VERSION : 0.1
   VAR
      General : Struct
         ManipulatorFaultProximitiSwitch : Bool;
         ManipulatorFaultRuntime : Bool;
         CPCleanerFaultProximitiSwitch : Bool;
         CPCleanerFaultRuntime : Bool;
         PCPCleaner : Bool;
         Spare6 : Bool;
         Spare7 : Bool;
         Spare8 : Bool;
         Spare9 : Bool;
         Spare10 : Bool;
         Spare11 : Bool;
         Spare12 : Bool;
         Spare13 : Bool;
         Spare14 : Bool;
         Spare15 : Bool;
         Spare16 : Bool;
      END_STRUCT;
      SafteyDeviceSelected : Array[1..16] of Bool;
      "Saftey DeviceAS" : Array[1..16] of Bool;   // Automatic stop at the Saftey Device
      "Saftey DeviceES" : Array[1..16] of Bool;   // Emergency stop at the Saftey Device
   END_VAR
BEGIN
END_DATA_BLOCK

DATA_BLOCK "DB1031_AddStatus"   // DB1031
{ S7_Optimized_Access := 'FALSE' }
VERSION : 0.1
   VAR
      SaftyDevice : Array[0..4] of "UDT_SafetyDevice";
   END_VAR
BEGIN
END_DATA_BLOCK

DATA_BLOCK "DB1040_TT_MovementFault"   // DB1040
{ S7_Optimized_Access := 'FALSE' }
VERSION : 0.1
   VAR
      General : Struct
         MLD_Taktdehnung1Aktiv : Bool;   // Taktdehnung 01 ist aktiv
         MLD_Taktdehnung2Aktiv : Bool;   // Taktdehnung 02 ist aktiv
         MLD_Taktdehnung3Aktiv : Bool;   // Taktdehnung 03 ist aktiv
         MLD_Taktdehnung4Aktiv : Bool;   // Taktdehnung 04 ist aktiv
         STG_Reserve_0_4 : Bool;
         STG_Reserve_0_5 : Bool;
         STG_Reserve_0_6 : Bool;
         STG_Reserve_0_7 : Bool;
         STG_Reserve_1_0 : Bool;
         STG_Reserve_1_1 : Bool;
         STG_Reserve_1_2 : Bool;
         STG_Reserve_1_3 : Bool;
         STG_Reserve_1_4 : Bool;
         STG_Reserve_1_5 : Bool;
         STG_Reserve_1_6 : Bool;
         STG_Reserve_1_7 : Bool;
      END_STRUCT;
      IPOS : Struct
         STG_Luefter : Bool;   // Störung Grp2: Der Versorgung oder des Motorschutzes des Lüfters
         STG_Umrichter : Bool;   // Störung: Der Umrichter ist nicht betriebsbereit
         STG_Motorschutz : Bool;   // Störung: Der Versorgung oder des Motorschutzes des Umrichters
         STG_von_IPOS : Bool;   // Störung: Ein Störungssignal von dem Umrichter steht an
         STG_Genauhaltini : Bool;   // Störung: Die Genauhalteposition (Initiator) wurde nicht erreicht
         STG_Genauhalt_immer_ein : Bool;   // Störung: Die Genauhalteposition (Initiator) wird dauernd belegt
         STG_Busfehler : Bool;   // Störung: Busteilnehmer ist nicht erreichbar
         STG_Reserve_0_7 : Bool;
         STG_Reserve_1_0 : Bool;
         STG_Reserve_1_1 : Bool;
         STG_Reserve_1_2 : Bool;
         STG_Reserve_1_3 : Bool;
         STG_Reserve_1_4 : Bool;
         STG_Reserve_1_5 : Bool;
         STG_Reserve_1_6 : Bool;
         STG_Reserve_1_7 : Bool;
      END_STRUCT;
      Segmentkennung : Struct
         STG_Nummer_unlogisch : Bool;
         STG_Hardwareabschaltung : Bool;
         STG_Wechsel_in_Pos : Bool;
         STG_Reserve_0_3 : Bool;
         STG_Reserve_0_4 : Bool;
         STG_Reserve_0_5 : Bool;
         STG_Reserve_0_6 : Bool;
         STG_Reserve_0_7 : Bool;
         STG_Reserve_1_0 : Bool;
         STG_Reserve_1_1 : Bool;
         STG_Reserve_1_2 : Bool;
         STG_Reserve_1_3 : Bool;
         STG_Reserve_1_4 : Bool;
         STG_Reserve_1_5 : Bool;
         STG_Reserve_1_6 : Bool;
         STG_Reserve_1_7 : Bool;
      END_STRUCT;
      Kettenspanner : Struct
         STG_Entlastung : Bool;
         STG_Druckaufbau : Bool;
         STG_Reserve_0_2 : Bool;
         STG_Reserve_0_3 : Bool;
         STG_Reserve_0_4 : Bool;
         STG_Reserve_0_5 : Bool;
         STG_Reserve_0_6 : Bool;
         STG_Reserve_0_7 : Bool;
         STG_Reserve_1_0 : Bool;
         STG_Reserve_1_1 : Bool;
         STG_Reserve_1_2 : Bool;
         STG_Reserve_1_3 : Bool;
         STG_Reserve_1_4 : Bool;
         STG_Reserve_1_5 : Bool;
         STG_Reserve_1_6 : Bool;
         STG_Reserve_1_7 : Bool;
      END_STRUCT;
   END_VAR
BEGIN
END_DATA_BLOCK

DATA_BLOCK "DB1049_TT_Value"   // DB1049
{ S7_Optimized_Access := 'FALSE' }
AUTHOR : KT242
VERSION : 0.1
   VAR
      Taktzeit : S5Time := S5T#15S;
      Vorwarnzeit : S5Time := S5T#1S;
      Seg_fuer_WW : Int := 0;
      Seg_fuer_Teachen : Int := 0;
      Pos_Offset_Stop : Int := 0;
      Pos_Offset_WW : Int := 0;
      Pos_Offset_Teachen : Int := 0;
      Antrieb_RP : Int := 5000;
      Antrieb_RN : Int := 5000;
      Antrieb_Hand : Int := 500;
      Antrieb_Auto : Int := 1200;
      WaitTimeMHFront : S5Time := S5T#2S;
      RunTimeManipulator : S5Time := S5T#30S;
      RunTimeCPCleaner : S5Time := S5T#5S;
      DelayTimeCPCleaning : S5Time := S5T#500MS;
      DurationCPCleaning : S5Time := S5T#2S;
   END_VAR
BEGIN
END_DATA_BLOCK

DATA_BLOCK "DB1050_Seg_Fault"   // DB1050
{ S7_Optimized_Access := 'FALSE' }
VERSION : 0.1
   VAR
      General : Struct
         STG_Reserve_0_0 : Bool;
         STG_Reserve_0_1 : Bool;
         STG_Reserve_0_2 : Bool;
         STG_Reserve_0_3 : Bool;
         STG_Reserve_0_4 : Bool;
         STG_Reserve_0_5 : Bool;
         STG_Reserve_0_6 : Bool;
         STG_Reserve_0_7 : Bool;
         STG_Reserve_1_0 : Bool;
         STG_Reserve_1_1 : Bool;
         STG_Reserve_1_2 : Bool;
         STG_Reserve_1_3 : Bool;
         STG_Reserve_1_4 : Bool;
         STG_Reserve_1_5 : Bool;
         STG_Reserve_1_6 : Bool;
         STG_Reserve_1_7 : Bool;
      END_STRUCT;
      Segmentverwaltung : Struct
         STG_keine_SegmentNr : Bool;   // Störung Grp3: Es ist keine Segmentkennung vorhanden
         STG_falsche_Paritaet : Bool;   // Störung Grp1: Das Paritätsbit wurde falsch gesetzt
         STG_SegNr_zu_gross : Bool;   // Störung Grp1: Die verdrahtete Segmentnummer ist für dieses RT zu Groß
         STG_Platz_doppelt : Bool;   // Störung Grp1: der Platz auf dem Segment wurde doppelt belegt // Verdrahtungsfehler
         STG_Reserve_0_4 : Bool;
         STG_Reserve_0_5 : Bool;
         STG_Reserve_0_6 : Bool;
         STG_Reserve_0_7 : Bool;
         STG_Reserve_1_0 : Bool;
         STG_Reserve_1_1 : Bool;
         STG_Reserve_1_2 : Bool;
         STG_Reserve_1_3 : Bool;
         STG_Reserve_1_4 : Bool;
         STG_Reserve_1_5 : Bool;
         STG_Reserve_1_6 : Bool;
         STG_Reserve_1_7 : Bool;
      END_STRUCT;
   END_VAR
BEGIN
END_DATA_BLOCK

DATA_BLOCK "DB1051_TT_SegValue"   // DB1051
{ S7_Optimized_Access := 'FALSE' }
VERSION : 0.1
   VAR
      Station : Array[1..8] of Struct
         FoamingEnable : Bool;
         MovingEnable : Bool;
         ToolChange : Bool;
         Spare4 : Bool;
         Spare5 : Bool;
         Spare6 : Bool;
         Spare7 : Bool;
         Spare8 : Bool;
         Spare9 : Bool;
         Spare10 : Bool;
         Spare11 : Bool;
         Spare12 : Bool;
         Spare13 : Bool;
         Spare14 : Bool;
         Spare15 : Bool;
         Spare16 : Bool;
         FoamingProg : Int;
         RobotProg : Int;
      END_STRUCT;
   END_VAR
BEGIN
   Station[1].FoamingEnable := TRUE;
   Station[1].MovingEnable := FALSE;
   Station[1].ToolChange := FALSE;
   Station[1].Spare4 := FALSE;
   Station[1].Spare5 := FALSE;
   Station[1].Spare6 := FALSE;
   Station[1].Spare7 := FALSE;
   Station[1].Spare8 := FALSE;
   Station[1].Spare9 := FALSE;
   Station[1].Spare10 := FALSE;
   Station[1].Spare11 := FALSE;
   Station[1].Spare12 := FALSE;
   Station[1].Spare13 := FALSE;
   Station[1].Spare14 := FALSE;
   Station[1].Spare15 := FALSE;
   Station[1].Spare16 := FALSE;
   Station[1].FoamingProg := 11;
   Station[1].RobotProg := 0;
   Station[2].FoamingEnable := FALSE;
   Station[2].MovingEnable := FALSE;
   Station[2].ToolChange := FALSE;
   Station[2].Spare4 := FALSE;
   Station[2].Spare5 := FALSE;
   Station[2].Spare6 := FALSE;
   Station[2].Spare7 := FALSE;
   Station[2].Spare8 := FALSE;
   Station[2].Spare9 := FALSE;
   Station[2].Spare10 := FALSE;
   Station[2].Spare11 := FALSE;
   Station[2].Spare12 := FALSE;
   Station[2].Spare13 := FALSE;
   Station[2].Spare14 := FALSE;
   Station[2].Spare15 := FALSE;
   Station[2].Spare16 := FALSE;
   Station[2].FoamingProg := 1;
   Station[2].RobotProg := 0;
   Station[3].FoamingEnable := FALSE;
   Station[3].MovingEnable := FALSE;
   Station[3].ToolChange := FALSE;
   Station[3].Spare4 := FALSE;
   Station[3].Spare5 := FALSE;
   Station[3].Spare6 := FALSE;
   Station[3].Spare7 := FALSE;
   Station[3].Spare8 := FALSE;
   Station[3].Spare9 := FALSE;
   Station[3].Spare10 := FALSE;
   Station[3].Spare11 := FALSE;
   Station[3].Spare12 := FALSE;
   Station[3].Spare13 := FALSE;
   Station[3].Spare14 := FALSE;
   Station[3].Spare15 := FALSE;
   Station[3].Spare16 := FALSE;
   Station[3].FoamingProg := 3;
   Station[3].RobotProg := 0;
   Station[4].FoamingEnable := TRUE;
   Station[4].MovingEnable := FALSE;
   Station[4].ToolChange := FALSE;
   Station[4].Spare4 := FALSE;
   Station[4].Spare5 := FALSE;
   Station[4].Spare6 := FALSE;
   Station[4].Spare7 := FALSE;
   Station[4].Spare8 := FALSE;
   Station[4].Spare9 := FALSE;
   Station[4].Spare10 := FALSE;
   Station[4].Spare11 := FALSE;
   Station[4].Spare12 := FALSE;
   Station[4].Spare13 := FALSE;
   Station[4].Spare14 := FALSE;
   Station[4].Spare15 := FALSE;
   Station[4].Spare16 := FALSE;
   Station[4].FoamingProg := 4;
   Station[4].RobotProg := 0;
   Station[5].FoamingEnable := FALSE;
   Station[5].MovingEnable := FALSE;
   Station[5].ToolChange := FALSE;
   Station[5].Spare4 := FALSE;
   Station[5].Spare5 := FALSE;
   Station[5].Spare6 := FALSE;
   Station[5].Spare7 := FALSE;
   Station[5].Spare8 := FALSE;
   Station[5].Spare9 := FALSE;
   Station[5].Spare10 := FALSE;
   Station[5].Spare11 := FALSE;
   Station[5].Spare12 := FALSE;
   Station[5].Spare13 := FALSE;
   Station[5].Spare14 := FALSE;
   Station[5].Spare15 := FALSE;
   Station[5].Spare16 := FALSE;
   Station[5].FoamingProg := 5;
   Station[5].RobotProg := 0;
   Station[6].FoamingEnable := TRUE;
   Station[6].MovingEnable := FALSE;
   Station[6].ToolChange := FALSE;
   Station[6].Spare4 := FALSE;
   Station[6].Spare5 := FALSE;
   Station[6].Spare6 := FALSE;
   Station[6].Spare7 := FALSE;
   Station[6].Spare8 := FALSE;
   Station[6].Spare9 := FALSE;
   Station[6].Spare10 := FALSE;
   Station[6].Spare11 := FALSE;
   Station[6].Spare12 := FALSE;
   Station[6].Spare13 := FALSE;
   Station[6].Spare14 := FALSE;
   Station[6].Spare15 := FALSE;
   Station[6].Spare16 := FALSE;
   Station[6].FoamingProg := 1;
   Station[6].RobotProg := 0;
   Station[7].FoamingEnable := FALSE;
   Station[7].MovingEnable := FALSE;
   Station[7].ToolChange := FALSE;
   Station[7].Spare4 := FALSE;
   Station[7].Spare5 := FALSE;
   Station[7].Spare6 := FALSE;
   Station[7].Spare7 := FALSE;
   Station[7].Spare8 := FALSE;
   Station[7].Spare9 := FALSE;
   Station[7].Spare10 := FALSE;
   Station[7].Spare11 := FALSE;
   Station[7].Spare12 := FALSE;
   Station[7].Spare13 := FALSE;
   Station[7].Spare14 := FALSE;
   Station[7].Spare15 := FALSE;
   Station[7].Spare16 := FALSE;
   Station[7].FoamingProg := 7;
   Station[7].RobotProg := 0;
   Station[8].FoamingEnable := FALSE;
   Station[8].MovingEnable := FALSE;
   Station[8].ToolChange := FALSE;
   Station[8].Spare4 := FALSE;
   Station[8].Spare5 := FALSE;
   Station[8].Spare6 := FALSE;
   Station[8].Spare7 := FALSE;
   Station[8].Spare8 := FALSE;
   Station[8].Spare9 := FALSE;
   Station[8].Spare10 := FALSE;
   Station[8].Spare11 := FALSE;
   Station[8].Spare12 := FALSE;
   Station[8].Spare13 := FALSE;
   Station[8].Spare14 := FALSE;
   Station[8].Spare15 := FALSE;
   Station[8].Spare16 := FALSE;
   Station[8].FoamingProg := 11;
   Station[8].RobotProg := 0;
END_DATA_BLOCK

DATA_BLOCK "DB1059_TTSegmentFault"   // DB1059
{ S7_Optimized_Access := 'FALSE' }
VERSION : 0.1
   VAR
      Bits : Struct
         Emptying : Bool;
         PressureSwitchNotreached : Bool;
         ProxySwitchNotReached : Bool;
      END_STRUCT;
      MouldNotExist : Array[1..16] of Bool;
      MouldNotClosed : Array[1..16] of Bool;
      MouldNoFoaming : Array[1..16] of Bool;
   END_VAR
BEGIN
END_DATA_BLOCK

DATA_BLOCK "DB1200_ProCanConf"   // DB1200
TITLE = Address allocation IO-ProCan
{ S7_Optimized_Access := 'FALSE' }
VERSION : 0.1
   VAR
      ReadWriteDeviceNo : Int := 1;
      CopyDeviceNO : Int := 0;
      Read : Bool := FALSE;
      Write : Bool := FALSE;
      Copy : Bool := FALSE;
      ProCanConf : Array[0..13] of "UDT1201_ProCanAddress";   // 1-4 Maschinenmodule; 5-36 Mischkopfmodule
   END_VAR
BEGIN
   ProCanConf[1].Output.Telegram_Recive := 1100;
   ProCanConf[1].Input.Telegram_Reserve := 0;
   ProCanConf[1].Flag_Modul_OK := TRUE;
   ProCanConf[1].Input.Telegram := 1100;
   ProCanConf[1].Address.MachineNo := 1;
   ProCanConf[1].Address.FlowNo01 := 1;
   ProCanConf[1].Address.FlowNo02 := 2;
   ProCanConf[1].Flag_Modul_NOK := TRUE;
   ProCanConf[2].Input.Telegram := 1100;
   ProCanConf[2].Output.Telegram_Recive := 1200;
   ProCanConf[2].Address.MixingheadNo01 := 1;
   ProCanConf[3].Input.Telegram := 1300;
   ProCanConf[3].Output.Telegram_Recive := 1300;
   ProCanConf[3].Address.MixingheadNo01 := 2;
   ProCanConf[4].Input.Telegram := 1400;
   ProCanConf[4].Output.Telegram_Recive := 1400;
   ProCanConf[4].Address.MixingheadNo01 := 3;
   ProCanConf[0].Input.Telegram := 1100;
   ProCanConf[0].Input.Telegram_Reserve := 0;
   ProCanConf[0].Output.Reserve01 := 0;
   ProCanConf[0].Output.Telegram_Recive := 1100;
   ProCanConf[0].Address.MachineNo := 1;
   ProCanConf[0].Address.FlowNo01 := 1;
   ProCanConf[0].Address.FlowNo02 := 2;
   ProCanConf[0].Address.FlowNo03 := 0;
   ProCanConf[0].Address.FlowNo04 := 0;
   ProCanConf[0].Address.MixingheadNo01 := 0;
   ProCanConf[0].Address.MixingheadNo02 := 0;
   ProCanConf[0].Address.BypassNozzelNo01 := 0;
   ProCanConf[0].Address.BypassNozzelNo02 := 0;
   ProCanConf[0].Address.MeteringPistonNo01 := 0;
   ProCanConf[0].Address.MeteringPistonNo02 := 0;
   ProCanConf[0].Address.MeteringPistonNo03 := 0;
   ProCanConf[0].Address.MeteringPistonNo04 := 0;
   ProCanConf[0].Address.TandemNo01 := 0;
   ProCanConf[0].Address.TandemNo02 := 0;
   ProCanConf[0].Address.PLC_No01 := 0;
   ProCanConf[0].Address.PLC_No02 := 0;
   ProCanConf[0].Address.PLC_No03 := 0;
   ProCanConf[0].Address.PLC_No04 := 0;
   ProCanConf[0].Flag_Modul_OK := TRUE;
   ProCanConf[0].Flag_Modul_NOK := TRUE;
   ProCanConf[0].Spare_02 := FALSE;
   ProCanConf[0].Spare_03 := FALSE;
   ProCanConf[0].Spare_04 := FALSE;
   ProCanConf[0].Spare_05 := FALSE;
   ProCanConf[0].Spare_06 := FALSE;
   ProCanConf[0].Spare_07 := FALSE;
   ProCanConf[0].Spare_08 := FALSE;
   ProCanConf[0].Spare_09 := FALSE;
   ProCanConf[0].Spare_010 := FALSE;
   ProCanConf[0].Spare_011 := FALSE;
   ProCanConf[0].Spare_012 := FALSE;
   ProCanConf[0].Spare_013 := FALSE;
   ProCanConf[0].Spare_014 := FALSE;
   ProCanConf[0].Spare_015 := FALSE;
   ProCanConf[1].Output.Reserve01 := 0;
   ProCanConf[1].Address.FlowNo03 := 0;
   ProCanConf[1].Address.FlowNo04 := 0;
   ProCanConf[1].Address.MixingheadNo01 := 0;
   ProCanConf[1].Address.MixingheadNo02 := 0;
   ProCanConf[1].Address.BypassNozzelNo01 := 0;
   ProCanConf[1].Address.BypassNozzelNo02 := 0;
   ProCanConf[1].Address.MeteringPistonNo01 := 0;
   ProCanConf[1].Address.MeteringPistonNo02 := 0;
   ProCanConf[1].Address.MeteringPistonNo03 := 0;
   ProCanConf[1].Address.MeteringPistonNo04 := 0;
   ProCanConf[1].Address.TandemNo01 := 0;
   ProCanConf[1].Address.TandemNo02 := 0;
   ProCanConf[1].Address.PLC_No01 := 0;
   ProCanConf[1].Address.PLC_No02 := 0;
   ProCanConf[1].Address.PLC_No03 := 0;
   ProCanConf[1].Address.PLC_No04 := 0;
   ProCanConf[1].Spare_02 := FALSE;
   ProCanConf[1].Spare_03 := FALSE;
   ProCanConf[1].Spare_04 := FALSE;
   ProCanConf[1].Spare_05 := FALSE;
   ProCanConf[1].Spare_06 := FALSE;
   ProCanConf[1].Spare_07 := FALSE;
   ProCanConf[1].Spare_08 := FALSE;
   ProCanConf[1].Spare_09 := FALSE;
   ProCanConf[1].Spare_010 := FALSE;
   ProCanConf[1].Spare_011 := FALSE;
   ProCanConf[1].Spare_012 := FALSE;
   ProCanConf[1].Spare_013 := FALSE;
   ProCanConf[1].Spare_014 := FALSE;
   ProCanConf[1].Spare_015 := FALSE;
   ProCanConf[2].Input.Telegram_Reserve := 0;
   ProCanConf[2].Output.Reserve01 := 0;
   ProCanConf[2].Address.MachineNo := 1;
   ProCanConf[2].Address.FlowNo01 := 0;
   ProCanConf[2].Address.FlowNo02 := 0;
   ProCanConf[2].Address.FlowNo03 := 0;
   ProCanConf[2].Address.FlowNo04 := 0;
   ProCanConf[2].Address.MixingheadNo02 := 0;
   ProCanConf[2].Address.BypassNozzelNo01 := 0;
   ProCanConf[2].Address.BypassNozzelNo02 := 0;
   ProCanConf[2].Address.MeteringPistonNo01 := 0;
   ProCanConf[2].Address.MeteringPistonNo02 := 0;
   ProCanConf[2].Address.MeteringPistonNo03 := 0;
   ProCanConf[2].Address.MeteringPistonNo04 := 0;
   ProCanConf[2].Address.TandemNo01 := 0;
   ProCanConf[2].Address.TandemNo02 := 0;
   ProCanConf[2].Address.PLC_No01 := 0;
   ProCanConf[2].Address.PLC_No02 := 0;
   ProCanConf[2].Address.PLC_No03 := 0;
   ProCanConf[2].Address.PLC_No04 := 0;
   ProCanConf[2].Flag_Modul_OK := TRUE;
   ProCanConf[2].Flag_Modul_NOK := TRUE;
   ProCanConf[2].Spare_02 := FALSE;
   ProCanConf[2].Spare_03 := FALSE;
   ProCanConf[2].Spare_04 := FALSE;
   ProCanConf[2].Spare_05 := FALSE;
   ProCanConf[2].Spare_06 := FALSE;
   ProCanConf[2].Spare_07 := FALSE;
   ProCanConf[2].Spare_08 := FALSE;
   ProCanConf[2].Spare_09 := FALSE;
   ProCanConf[2].Spare_010 := FALSE;
   ProCanConf[2].Spare_011 := FALSE;
   ProCanConf[2].Spare_012 := FALSE;
   ProCanConf[2].Spare_013 := FALSE;
   ProCanConf[2].Spare_014 := FALSE;
   ProCanConf[2].Spare_015 := FALSE;
   ProCanConf[3].Input.Telegram_Reserve := 0;
   ProCanConf[3].Output.Reserve01 := 0;
   ProCanConf[3].Address.MachineNo := 0;
   ProCanConf[3].Address.FlowNo01 := 4;
   ProCanConf[3].Address.FlowNo02 := 0;
   ProCanConf[3].Address.FlowNo03 := 0;
   ProCanConf[3].Address.FlowNo04 := 0;
   ProCanConf[3].Address.MixingheadNo02 := 0;
   ProCanConf[3].Address.BypassNozzelNo01 := 0;
   ProCanConf[3].Address.BypassNozzelNo02 := 0;
   ProCanConf[3].Address.MeteringPistonNo01 := 0;
   ProCanConf[3].Address.MeteringPistonNo02 := 0;
   ProCanConf[3].Address.MeteringPistonNo03 := 0;
   ProCanConf[3].Address.MeteringPistonNo04 := 0;
   ProCanConf[3].Address.TandemNo01 := 0;
   ProCanConf[3].Address.TandemNo02 := 0;
   ProCanConf[3].Address.PLC_No01 := 0;
   ProCanConf[3].Address.PLC_No02 := 0;
   ProCanConf[3].Address.PLC_No03 := 0;
   ProCanConf[3].Address.PLC_No04 := 0;
   ProCanConf[3].Flag_Modul_OK := FALSE;
   ProCanConf[3].Flag_Modul_NOK := FALSE;
   ProCanConf[3].Spare_02 := FALSE;
   ProCanConf[3].Spare_03 := FALSE;
   ProCanConf[3].Spare_04 := FALSE;
   ProCanConf[3].Spare_05 := FALSE;
   ProCanConf[3].Spare_06 := FALSE;
   ProCanConf[3].Spare_07 := FALSE;
   ProCanConf[3].Spare_08 := FALSE;
   ProCanConf[3].Spare_09 := FALSE;
   ProCanConf[3].Spare_010 := FALSE;
   ProCanConf[3].Spare_011 := FALSE;
   ProCanConf[3].Spare_012 := FALSE;
   ProCanConf[3].Spare_013 := FALSE;
   ProCanConf[3].Spare_014 := FALSE;
   ProCanConf[3].Spare_015 := FALSE;
   ProCanConf[4].Input.Telegram_Reserve := 0;
   ProCanConf[4].Output.Reserve01 := 0;
   ProCanConf[4].Address.MachineNo := 0;
   ProCanConf[4].Address.FlowNo01 := 5;
   ProCanConf[4].Address.FlowNo02 := 0;
   ProCanConf[4].Address.FlowNo03 := 0;
   ProCanConf[4].Address.FlowNo04 := 0;
   ProCanConf[4].Address.MixingheadNo02 := 0;
   ProCanConf[4].Address.BypassNozzelNo01 := 0;
   ProCanConf[4].Address.BypassNozzelNo02 := 0;
   ProCanConf[4].Address.MeteringPistonNo01 := 0;
   ProCanConf[4].Address.MeteringPistonNo02 := 0;
   ProCanConf[4].Address.MeteringPistonNo03 := 0;
   ProCanConf[4].Address.MeteringPistonNo04 := 0;
   ProCanConf[4].Address.TandemNo01 := 0;
   ProCanConf[4].Address.TandemNo02 := 0;
   ProCanConf[4].Address.PLC_No01 := 0;
   ProCanConf[4].Address.PLC_No02 := 0;
   ProCanConf[4].Address.PLC_No03 := 0;
   ProCanConf[4].Address.PLC_No04 := 0;
   ProCanConf[4].Flag_Modul_OK := FALSE;
   ProCanConf[4].Flag_Modul_NOK := FALSE;
   ProCanConf[4].Spare_02 := FALSE;
   ProCanConf[4].Spare_03 := FALSE;
   ProCanConf[4].Spare_04 := FALSE;
   ProCanConf[4].Spare_05 := FALSE;
   ProCanConf[4].Spare_06 := FALSE;
   ProCanConf[4].Spare_07 := FALSE;
   ProCanConf[4].Spare_08 := FALSE;
   ProCanConf[4].Spare_09 := FALSE;
   ProCanConf[4].Spare_010 := FALSE;
   ProCanConf[4].Spare_011 := FALSE;
   ProCanConf[4].Spare_012 := FALSE;
   ProCanConf[4].Spare_013 := FALSE;
   ProCanConf[4].Spare_014 := FALSE;
   ProCanConf[4].Spare_015 := FALSE;
   ProCanConf[5].Input.Telegram := 1500;
   ProCanConf[5].Input.Telegram_Reserve := 0;
   ProCanConf[5].Output.Reserve01 := 0;
   ProCanConf[5].Output.Telegram_Recive := 1500;
   ProCanConf[5].Address.MachineNo := 0;
   // 346 more start values not shown
END_DATA_BLOCK

DATA_BLOCK "DB1232_ProCanIO_MH"   // DB1232
TITLE = Address allocation mixing head IO-ProCan
{ S7_Optimized_Access := 'FALSE' }
VERSION : 0.1
   VAR
      ReadWriteDeviceNo : Int := 1;
      CopyDeviceNO : Int := 0;
      Read : Bool := FALSE;
      Write : Bool := FALSE;
      Copy : Bool := FALSE;
      AddressMH : Array[0..16] of "UDT1232_ProCanIO_MH";
   END_VAR
BEGIN
   AddressMH[1].Ref_Digital_Input := 20;
   AddressMH[1].Ref_MH_ShotTime := 1250;
   AddressMH[1].Ref_MH_Opening_Time := 1254;
   AddressMH[1].Ref_MH_Closing_Time := 1256;
   AddressMH[1].Ref_MH_State := 1260;
   AddressMH[1].Ref_Digital_Output := 20;
   AddressMH[1].Ref_ShotTimeSetValue := 1250;
   AddressMH[1].Ref_ServiceProduction := 1254;
   AddressMH[1].Ref_MixingheadControl := 1260;
   AddressMH[1].Ref_OK := TRUE;
   AddressMH[1].MH_Channel_01 := TRUE;
   AddressMH[2].Ref_Digital_Input := 24;
   AddressMH[2].Ref_MH_ShotTime := 1350;
   AddressMH[2].Ref_MH_Opening_Time := 1354;
   AddressMH[2].Ref_MH_Closing_Time := 1356;
   AddressMH[2].Ref_MH_State := 1360;
   AddressMH[2].Ref_Digital_Output := 24;
   AddressMH[2].Ref_ShotTimeSetValue := 1350;
   AddressMH[2].Ref_ServiceProduction := 1354;
   AddressMH[2].Ref_MixingheadControl := 1360;
   AddressMH[3].Ref_Digital_Input := 28;
   AddressMH[3].Ref_MH_ShotTime := 1450;
   AddressMH[3].Ref_MH_Opening_Time := 1454;
   AddressMH[3].Ref_MH_Closing_Time := 1456;
   AddressMH[3].Ref_MH_State := 1460;
   AddressMH[3].Ref_Digital_Output := 28;
   AddressMH[3].Ref_ShotTimeSetValue := 1450;
   AddressMH[3].Ref_ServiceProduction := 1454;
   AddressMH[3].Ref_MixingheadControl := 1460;
   AddressMH[0].Ref_Digital_Input := 20;
   AddressMH[0].Ref_MH_ShotTime := 1250;
   AddressMH[0].Ref_MH_Opening_Time := 1254;
   AddressMH[0].Ref_MH_Closing_Time := 1256;
   AddressMH[0].Ref_MH_State := 1260;
   AddressMH[0].Ref_PLC_State := 0;
   AddressMH[0].Ref_CP_State := 0;
   AddressMH[0].Ref_Digital_Output := 20;
   AddressMH[0].Ref_ShotTimeSetValue := 1250;
   AddressMH[0].Ref_ServiceProduction := 1254;
   AddressMH[0].Ref_MixingheadControl := 1260;
   AddressMH[0].Ref_PLC_comand_SP := 0;
   AddressMH[0].Ref_PLC_comand_CP := 0;
   AddressMH[0].Ref_PLC_set_value_SP := 0;
   AddressMH[0].Ref_PLC_set_value_CP := 0;
   AddressMH[0].Ref_NozzelBypassControl := 0;
   AddressMH[0].Ref_NozzelBypassSetOut := 0;
   AddressMH[0].Ref_Reserve := 0;
   AddressMH[0].Ref_OK := TRUE;
   AddressMH[0].MH_Channel_01 := TRUE;
   AddressMH[0].MH_Channel_02 := FALSE;
   AddressMH[0].Spare_03 := FALSE;
   AddressMH[0].Spare_04 := FALSE;
   AddressMH[0].Spare_05 := FALSE;
   AddressMH[0].Spare_06 := FALSE;
   AddressMH[0].Spare_07 := FALSE;
   AddressMH[1].Ref_PLC_State := 0;
   AddressMH[1].Ref_CP_State := 0;
   AddressMH[1].Ref_PLC_comand_SP := 0;
   AddressMH[1].Ref_PLC_comand_CP := 0;
   AddressMH[1].Ref_PLC_set_value_SP := 0;
   AddressMH[1].Ref_PLC_set_value_CP := 0;
   AddressMH[1].Ref_NozzelBypassControl := 0;
   AddressMH[1].Ref_NozzelBypassSetOut := 0;
   AddressMH[1].Ref_Reserve := 0;
   AddressMH[1].MH_Channel_02 := FALSE;
   AddressMH[1].Spare_03 := FALSE;
   AddressMH[1].Spare_04 := FALSE;
   AddressMH[1].Spare_05 := FALSE;
   AddressMH[1].Spare_06 := FALSE;
   AddressMH[1].Spare_07 := FALSE;
   AddressMH[2].Ref_PLC_State := 0;
   AddressMH[2].Ref_CP_State := 0;
   AddressMH[2].Ref_PLC_comand_SP := 0;
   AddressMH[2].Ref_PLC_comand_CP := 0;
   AddressMH[2].Ref_PLC_set_value_SP := 0;
   AddressMH[2].Ref_PLC_set_value_CP := 0;
   AddressMH[2].Ref_NozzelBypassControl := 0;
   AddressMH[2].Ref_NozzelBypassSetOut := 0;
   AddressMH[2].Ref_Reserve := 0;
   AddressMH[2].Ref_OK := FALSE;
   AddressMH[2].MH_Channel_01 := TRUE;
   AddressMH[2].MH_Channel_02 := FALSE;
   AddressMH[2].Spare_03 := FALSE;
   AddressMH[2].Spare_04 := FALSE;
   AddressMH[2].Spare_05 := FALSE;
   AddressMH[2].Spare_06 := FALSE;
   AddressMH[2].Spare_07 := FALSE;
   AddressMH[3].Ref_PLC_State := 0;
   AddressMH[3].Ref_CP_State := 0;
   AddressMH[3].Ref_PLC_comand_SP := 0;
   AddressMH[3].Ref_PLC_comand_CP := 0;
   AddressMH[3].Ref_PLC_set_value_SP := 0;